   "CARRIER #01 SpareSafetyOutput(3_2)" : Bool = PLC "CARRIER #01 SpareSafetyOutput(3_2)" AT %M84.1, 1 s
   "CARRIER #01 SpareSafetyOutput(3_3)" : Bool = PLC "CARRIER #01 SpareSafetyOutput(3_3)" AT %M84.2, 1 s
   "CARRIER #01 SpareSafetyOutput(3_4)" : Bool = PLC "CARRIER #01 SpareSafetyOutput(3_4)" AT %M84.3, 1 s
   "CARRIER #01 SpareSafetyOutput(3_5)" : Bool = PLC "CARRIER #01 SpareSafetyOutput(3_5)" AT %M84.4, 1 s
   "CARRIER #01 SpareSafetyOutput(3_6)" : Bool = PLC "CARRIER #01 SpareSafetyOutput(3_6)" AT %M84.5, 1 s
   "CARRIER #01 SpareSafetyOutput(3_7)" : Bool = PLC "CARRIER #01 SpareSafetyOutput(3_7)" AT %M84.6, 1 s
   "Carrier #01_ At Command Position" : Bool = PLC DB_SDC_ERRORS_STAT.ER_AKT[49].ER_STAT[1].ERROR AT %M84.7, 1 s
   "Carrier #01_ Carrier in zone" : Int = PLC "Carrier #01_ Carrier in zone" AT %MW86, 1 s
   "Carrier #01_ Next carrier number" : Int = PLC "Carrier #01_ Next carrier number" AT %MW88, 1 s
   "Carrier 1 G120 D Status" : Bool = PLC EMS.Carrier[12].SDC_IN.DriveCommFault AT %I412.1, 1 s
   "Carrier 1 HMI Status" : Bool = PLC "Carrier 1 HMI Status" AT %I412.2, 1 s
   "Carrier 1 PnF Encoder Status" : Bool = PLC "Carrier 1 PnF Encoder Status" AT %I412.0, 1 s
   "Carrier 2  HMI Staus" : Bool = PLC "Carrier 2 HMI Status" AT %I432.2, 1 s
   "Carrier 2 G120 D Status" : Bool = PLC "Carrier 2  Drive Status" AT %I432.1, 1 s
   "Carrier 2 PnF Encoder Status" : Bool = PLC "Carrier 2 PnF Encoder Status" AT %I432.0, 1 s
   "Carrier 3  G120 D Status" : Bool = PLC "Carrier 3  Drive Status" AT %I452.1, 1 s
   "Carrier 3  PnF Encoder Status" : Bool = PLC "Carrier 3 PnF Encoder Status" AT %I452.0, 1 s
   "Carrier 3 HMI Status" : Bool = PLC "Carrier 3 HMI Status" AT %I452.2, 1 s
   "Carrier 4 G120 D Status" : Bool = PLC "Carrier 4  Drive Status" AT %I472.1, 1 s
   "Carrier 4 HMI Status" : Bool = PLC "Carrier 4 HMI Status" AT %I472.2, 1 s
   "Carrier 4 PnF Encoder Status" : Bool = PLC "Carrier 4 PnF Encoder Status" AT %I472.0, 1 s
   "Carrier_Index_HMI" : Int = PLC Carrier_Index_HMI AT %MW70, 1 s
   "Always_OFF_HMI" : Bool, internal
   "Always_ON_HMI" : Bool, internal
   "EMS_Accum_Zone_Speed" : Word = PLC EMS.AccumZnSpeed AT %DB1.DBW0, 1 s
   "PLC_IP_Address" : WString[30], internal
   "DB302_HMI_Faults_Carrier1_Faults_0" : Int = PLC DB302_HMI_Faults.Carrier1_Faults_0 AT %DB1.DBW0, 1 s
   "DB302_HMI_Faults_Carrier1_Faults_1" : Int = PLC DB302_HMI_Faults.Carrier1_Faults_1 AT %DB1.DBW0, 1 s
   "DB302_HMI_Faults_Carrier1_Faults_2" : Int = PLC DB302_HMI_Faults.Carrier1_Faults_2 AT %DB1.DBW0, 1 s
   "DB302_HMI_Faults_Carrier1_Faults_3" : Int = PLC DB302_HMI_Faults.Carrier1_Faults_3 AT %DB1.DBW0, 1 s
   "DB302_HMI_Faults_Carrier10_Faults_0" : Int = PLC DB302_HMI_Faults.Carrier10_Faults_0 AT %DB1.DBW0, 1 s
   "DB302_HMI_Faults_Carrier10_Faults_1" : Int = PLC DB302_HMI_Faults.Carrier10_Faults_1 AT %DB1.DBW0, 1 s
   "DB302_HMI_Faults_Carrier10_Faults_2" : Int = PLC DB302_HMI_Faults.Carrier10_Faults_2 AT %DB1.DBW0, 1 s
   "DB302_HMI_Faults_Carrier10_Faults_3" : Int = PLC DB302_HMI_Faults.Carrier10_Faults_3 AT %DB1.DBW0, 1 s
   "DB302_HMI_Faults_Carrier11_Faults_0" : Int = PLC DB302_HMI_Faults.Carrier11_Faults_0 AT %DB1.DBW0, 1 s
   "DB302_HMI_Faults_Carrier11_Faults_1" : Int = PLC DB302_HMI_Faults.Carrier11_Faults_1 AT %DB1.DBW0, 1 s
   "DB302_HMI_Faults_Carrier11_Faults_2" : Int = PLC DB302_HMI_Faults.Carrier11_Faults_2 AT %DB1.DBW0, 1 s
   "DB302_HMI_Faults_Carrier11_Faults_3" : Int = PLC DB302_HMI_Faults.Carrier11_Faults_3 AT %DB1.DBW0, 1 s
   "DB302_HMI_Faults_Carrier12_Faults_0" : Int = PLC DB302_HMI_Faults.Carrier12_Faults_0 AT %DB1.DBW0, 1 s
   "DB302_HMI_Faults_Carrier12_Faults_1" : Int = PLC DB302_HMI_Faults.Carrier12_Faults_1 AT %DB1.DBW0, 1 s
   "DB302_HMI_Faults_Carrier12_Faults_2" : Int = PLC DB302_HMI_Faults.Carrier12_Faults_2 AT %DB1.DBW0, 1 s
   "DB302_HMI_Faults_Carrier12_Faults_3" : Int = PLC DB302_HMI_Faults.Carrier12_Faults_3 AT %DB1.DBW0, 1 s
   "DB302_HMI_Faults_Carrier13_Faults_0" : Int = PLC DB302_HMI_Faults.Carrier13_Faults_0 AT %DB1.DBW0, 1 s
   "DB302_HMI_Faults_Carrier13_Faults_1" : Int = PLC DB302_HMI_Faults.Carrier13_Faults_1 AT %DB1.DBW0, 1 s
   "DB302_HMI_Faults_Carrier13_Faults_2" : Int = PLC DB302_HMI_Faults.Carrier13_Faults_2 AT %DB1.DBW0, 1 s
   "DB302_HMI_Faults_Carrier13_Faults_3" : Int = PLC DB302_HMI_Faults.Carrier13_Faults_3 AT %DB1.DBW0, 1 s
   "DB302_HMI_Faults_Carrier14_Faults_0" : Int = PLC DB302_HMI_Faults.Carrier14_Faults_0 AT %DB1.DBW0, 1 s
   "DB302_HMI_Faults_Carrier14_Faults_1" : Int = PLC DB302_HMI_Faults.Carrier14_Faults_1 AT %DB1.DBW0, 1 s
   "DB302_HMI_Faults_Carrier14_Faults_2" : Int = PLC DB302_HMI_Faults.Carrier14_Faults_2 AT %DB1.DBW0, 1 s
   "DB302_HMI_Faults_Carrier14_Faults_3" : Int = PLC DB302_HMI_Faults.Carrier14_Faults_3 AT %DB1.DBW0, 1 s
   "DB302_HMI_Faults_Carrier15_Faults_0" : Int = PLC DB302_HMI_Faults.Carrier15_Faults_0 AT %DB1.DBW0, 1 s
   "DB302_HMI_Faults_Carrier15_Faults_1" : Int = PLC DB302_HMI_Faults.Carrier15_Faults_1 AT %DB1.DBW0, 1 s
   "DB302_HMI_Faults_Carrier15_Faults_2" : Int = PLC DB302_HMI_Faults.Carrier15_Faults_2 AT %DB1.DBW0, 1 s
   "DB302_HMI_Faults_Carrier15_Faults_3" : Int = PLC DB302_HMI_Faults.Carrier15_Faults_3 AT %DB1.DBW0, 1 s
   "DB302_HMI_Faults_Carrier16_Faults_0" : Int = PLC DB302_HMI_Faults.Carrier16_Faults_0 AT %DB1.DBW0, 1 s
   "DB302_HMI_Faults_Carrier16_Faults_1" : Int = PLC DB302_HMI_Faults.Carrier16_Faults_1 AT %DB1.DBW0, 1 s
   "DB302_HMI_Faults_Carrier16_Faults_2" : Int = PLC DB302_HMI_Faults.Carrier16_Faults_2 AT %DB1.DBW0, 1 s
   "DB302_HMI_Faults_Carrier16_Faults_3" : Int = PLC DB302_HMI_Faults.Carrier16_Faults_3 AT %DB1.DBW0, 1 s
   "DB302_HMI_Faults_Carrier17_Faults_0" : Int = PLC DB302_HMI_Faults.Carrier17_Faults_0 AT %DB1.DBW0, 1 s
   "DB302_HMI_Faults_Carrier17_Faults_1" : Int = PLC DB302_HMI_Faults.Carrier17_Faults_1 AT %DB1.DBW0, 1 s
   "DB302_HMI_Faults_Carrier17_Faults_2" : Int = PLC DB302_HMI_Faults.Carrier17_Faults_2 AT %DB1.DBW0, 1 s
   "DB302_HMI_Faults_Carrier17_Faults_3" : Int = PLC DB302_HMI_Faults.Carrier17_Faults_3 AT %DB1.DBW0, 1 s
   "DB302_HMI_Faults_Carrier18_Faults_0" : Int = PLC DB302_HMI_Faults.Carrier18_Faults_0 AT %DB1.DBW0, 1 s
   "DB302_HMI_Faults_Carrier18_Faults_1" : Int = PLC DB302_HMI_Faults.Carrier18_Faults_1 AT %DB1.DBW0, 1 s
   "DB302_HMI_Faults_Carrier18_Faults_2" : Int = PLC DB302_HMI_Faults.Carrier18_Faults_2 AT %DB1.DBW0, 1 s
   "DB302_HMI_Faults_Carrier18_Faults_3" : Int = PLC DB302_HMI_Faults.Carrier18_Faults_3 AT %DB1.DBW0, 1 s
   "DB302_HMI_Faults_Carrier19_Faults_0" : Int = PLC DB302_HMI_Faults.Carrier19_Faults_0 AT %DB1.DBW0, 1 s
   "DB302_HMI_Faults_Carrier19_Faults_1" : Int = PLC DB302_HMI_Faults.Carrier19_Faults_1 AT %DB1.DBW0, 1 s
   "DB302_HMI_Faults_Carrier19_Faults_2" : Int = PLC DB302_HMI_Faults.Carrier19_Faults_2 AT %DB1.DBW0, 1 s
   "DB302_HMI_Faults_Carrier19_Faults_3" : Int = PLC DB302_HMI_Faults.Carrier19_Faults_3 AT %DB1.DBW0, 1 s
   "DB302_HMI_Faults_Carrier2_Faults_0" : Int = PLC DB302_HMI_Faults.Carrier2_Faults_0 AT %DB1.DBW0, 1 s
   "DB302_HMI_Faults_Carrier2_Faults_1" : Int = PLC DB302_HMI_Faults.Carrier2_Faults_1 AT %DB1.DBW0, 1 s
   "DB302_HMI_Faults_Carrier2_Faults_2" : Int = PLC DB302_HMI_Faults.Carrier2_Faults_2 AT %DB1.DBW0, 1 s
   "DB302_HMI_Faults_Carrier2_Faults_3" : Int = PLC DB302_HMI_Faults.Carrier2_Faults_3 AT %DB1.DBW0, 1 s
   "DB302_HMI_Faults_Carrier20_Faults_0" : Int = PLC DB302_HMI_Faults.Carrier20_Faults_0 AT %DB1.DBW0, 1 s
   "DB302_HMI_Faults_Carrier20_Faults_1" : Int = PLC DB302_HMI_Faults.Carrier20_Faults_1 AT %DB1.DBW0, 1 s
   "DB302_HMI_Faults_Carrier20_Faults_2" : Int = PLC DB302_HMI_Faults.Carrier20_Faults_2 AT %DB1.DBW0, 1 s
   "DB302_HMI_Faults_Carrier20_Faults_3" : Int = PLC DB302_HMI_Faults.Carrier20_Faults_3 AT %DB1.DBW0, 1 s
   "DB302_HMI_Faults_Carrier21_Faults_0" : Int = PLC DB302_HMI_Faults.Carrier21_Faults_0 AT %DB1.DBW0, 1 s
   "DB302_HMI_Faults_Carrier21_Faults_1" : Int = PLC DB302_HMI_Faults.Carrier21_Faults_1 AT %DB1.DBW0, 1 s
   "DB302_HMI_Faults_Carrier21_Faults_2" : Int = PLC DB302_HMI_Faults.Carrier21_Faults_2 AT %DB1.DBW0, 1 s
   "DB302_HMI_Faults_Carrier21_Faults_3" : Int = PLC DB302_HMI_Faults.Carrier21_Faults_3 AT %DB1.DBW0, 1 s
   "DB302_HMI_Faults_Carrier22_Faults_0" : Int = PLC DB302_HMI_Faults.Carrier22_Faults_0 AT %DB1.DBW0, 1 s
   "DB302_HMI_Faults_Carrier22_Faults_1" : Int = PLC DB302_HMI_Faults.Carrier22_Faults_1 AT %DB1.DBW0, 1 s
   "DB302_HMI_Faults_Carrier22_Faults_2" : Int = PLC DB302_HMI_Faults.Carrier22_Faults_2 AT %DB1.DBW0, 1 s
   "DB302_HMI_Faults_Carrier22_Faults_3" : Int = PLC DB302_HMI_Faults.Carrier22_Faults_3 AT %DB1.DBW0, 1 s
   "DB302_HMI_Faults_Carrier23_Faults_0" : Int = PLC DB302_HMI_Faults.Carrier23_Faults_0 AT %DB1.DBW0, 1 s
   "DB302_HMI_Faults_Carrier23_Faults_1" : Int = PLC DB302_HMI_Faults.Carrier23_Faults_1 AT %DB1.DBW0, 1 s
   "DB302_HMI_Faults_Carrier23_Faults_2" : Int = PLC DB302_HMI_Faults.Carrier23_Faults_2 AT %DB1.DBW0, 1 s
   "DB302_HMI_Faults_Carrier23_Faults_3" : Int = PLC DB302_HMI_Faults.Carrier23_Faults_3 AT %DB1.DBW0, 1 s
   "DB302_HMI_Faults_Carrier24_Faults_0" : Int = PLC DB302_HMI_Faults.Carrier24_Faults_0 AT %DB1.DBW0, 1 s
   "DB302_HMI_Faults_Carrier24_Faults_1" : Int = PLC DB302_HMI_Faults.Carrier24_Faults_1 AT %DB1.DBW0, 1 s
   "DB302_HMI_Faults_Carrier24_Faults_2" : Int = PLC DB302_HMI_Faults.Carrier24_Faults_2 AT %DB1.DBW0, 1 s
   "DB302_HMI_Faults_Carrier24_Faults_3" : Int = PLC DB302_HMI_Faults.Carrier24_Faults_3 AT %DB1.DBW0, 1 s
   "DB302_HMI_Faults_Carrier25_Faults_0" : Int = PLC DB302_HMI_Faults.Carrier25_Faults_0 AT %DB1.DBW0, 1 s
   "DB302_HMI_Faults_Carrier25_Faults_1" : Int = PLC DB302_HMI_Faults.Carrier25_Faults_1 AT %DB1.DBW0, 1 s
   "DB302_HMI_Faults_Carrier25_Faults_2" : Int = PLC DB302_HMI_Faults.Carrier25_Faults_2 AT %DB1.DBW0, 1 s
   "DB302_HMI_Faults_Carrier25_Faults_3" : Int = PLC DB302_HMI_Faults.Carrier25_Faults_3 AT %DB1.DBW0, 1 s
   "DB302_HMI_Faults_Carrier26_Faults_0" : Int = PLC DB302_HMI_Faults.Carrier26_Faults_0 AT %DB1.DBW0, 1 s
   "DB302_HMI_Faults_Carrier26_Faults_1" : Int = PLC DB302_HMI_Faults.Carrier26_Faults_1 AT %DB1.DBW0, 1 s
   "DB302_HMI_Faults_Carrier26_Faults_2" : Int = PLC DB302_HMI_Faults.Carrier26_Faults_2 AT %DB1.DBW0, 1 s
   "DB302_HMI_Faults_Carrier26_Faults_3" : Int = PLC DB302_HMI_Faults.Carrier26_Faults_3 AT %DB1.DBW0, 1 s
   "DB302_HMI_Faults_Carrier27_Faults_0" : Int = PLC DB302_HMI_Faults.Carrier27_Faults_0 AT %DB1.DBW0, 1 s
   "DB302_HMI_Faults_Carrier27_Faults_1" : Int = PLC DB302_HMI_Faults.Carrier27_Faults_1 AT %DB1.DBW0, 1 s
   "DB302_HMI_Faults_Carrier27_Faults_2" : Int = PLC DB302_HMI_Faults.Carrier27_Faults_2 AT %DB1.DBW0, 1 s
   "DB302_HMI_Faults_Carrier27_Faults_3" : Int = PLC DB302_HMI_Faults.Carrier27_Faults_3 AT %DB1.DBW0, 1 s
   "DB302_HMI_Faults_Carrier28_Faults_0" : Int = PLC DB302_HMI_Faults.Carrier28_Faults_0 AT %DB1.DBW0, 1 s
   "DB302_HMI_Faults_Carrier28_Faults_1" : Int = PLC DB302_HMI_Faults.Carrier28_Faults_1 AT %DB1.DBW0, 1 s
   "DB302_HMI_Faults_Carrier28_Faults_2" : Int = PLC DB302_HMI_Faults.Carrier28_Faults_2 AT %DB1.DBW0, 1 s
   "DB302_HMI_Faults_Carrier28_Faults_3" : Int = PLC DB302_HMI_Faults.Carrier28_Faults_3 AT %DB1.DBW0, 1 s
   "DB302_HMI_Faults_Carrier29_Faults_0" : Int = PLC DB302_HMI_Faults.Carrier29_Faults_0 AT %DB1.DBW0, 1 s
   "DB302_HMI_Faults_Carrier29_Faults_1" : Int = PLC DB302_HMI_Faults.Carrier29_Faults_1 AT %DB1.DBW0, 1 s
   "DB302_HMI_Faults_Carrier29_Faults_2" : Int = PLC DB302_HMI_Faults.Carrier29_Faults_2 AT %DB1.DBW0, 1 s
   "DB302_HMI_Faults_Carrier29_Faults_3" : Int = PLC DB302_HMI_Faults.Carrier29_Faults_3 AT %DB1.DBW0, 1 s
   "DB302_HMI_Faults_Carrier3_Faults_0" : Int = PLC DB302_HMI_Faults.Carrier3_Faults_0 AT %DB1.DBW0, 1 s
   "DB302_HMI_Faults_Carrier3_Faults_1" : Int = PLC DB302_HMI_Faults.Carrier3_Faults_1 AT %DB1.DBW0, 1 s
   "DB302_HMI_Faults_Carrier3_Faults_2" : Int = PLC DB302_HMI_Faults.Carrier3_Faults_2 AT %DB1.DBW0, 1 s
   "DB302_HMI_Faults_Carrier3_Faults_3" : Int = PLC DB302_HMI_Faults.Carrier3_Faults_3 AT %DB1.DBW0, 1 s
   "DB302_HMI_Faults_Carrier30_Faults_0" : Int = PLC DB302_HMI_Faults.Carrier30_Faults_0 AT %DB1.DBW0, 1 s
   "DB302_HMI_Faults_Carrier30_Faults_1" : Int = PLC DB302_HMI_Faults.Carrier30_Faults_1 AT %DB1.DBW0, 1 s
   "DB302_HMI_Faults_Carrier30_Faults_2" : Int = PLC DB_SDC_ERRORS_STAT.ER_AKT[16].ER_STAT[2].DRIVE_POS AT %DB1.DBW0, 1 s
   "DB302_HMI_Faults_Carrier30_Faults_3" : Int = PLC DB302_HMI_Faults.Carrier30_Faults_3 AT %DB1.DBW0, 1 s
   "DB302_HMI_Faults_Carrier31_Faults_0" : Int = PLC DB302_HMI_Faults.Carrier31_Faults_0 AT %DB1.DBW0, 1 s
   "DB302_HMI_Faults_Carrier31_Faults_1" : Int = PLC DB302_HMI_Faults.Carrier31_Faults_1 AT %DB1.DBW0, 1 s
   "DB302_HMI_Faults_Carrier31_Faults_2" : Int = PLC DB302_HMI_Faults.Carrier31_Faults_2 AT %DB1.DBW0, 1 s
   "DB302_HMI_Faults_Carrier31_Faults_3" : Int = PLC DB302_HMI_Faults.Carrier31_Faults_3 AT %DB1.DBW0, 1 s
   "DB302_HMI_Faults_Carrier32_Faults_0" : Int = PLC DB302_HMI_Faults.Carrier32_Faults_0 AT %DB1.DBW0, 1 s
   "DB302_HMI_Faults_Carrier32_Faults_1" : Int = PLC DB302_HMI_Faults.Carrier32_Faults_1 AT %DB1.DBW0, 1 s
   "DB302_HMI_Faults_Carrier32_Faults_2" : Int = PLC DB302_HMI_Faults.Carrier32_Faults_2 AT %DB1.DBW0, 1 s
   "DB302_HMI_Faults_Carrier32_Faults_3" : Int = PLC DB302_HMI_Faults.Carrier32_Faults_3 AT %DB1.DBW0, 1 s
   "DB302_HMI_Faults_Carrier33_Faults_0" : Int = PLC DB302_HMI_Faults.Carrier33_Faults_0 AT %DB1.DBW0, 1 s
   "DB302_HMI_Faults_Carrier33_Faults_1" : Int = PLC DB302_HMI_Faults.Carrier33_Faults_1 AT %DB1.DBW0, 1 s
   "DB302_HMI_Faults_Carrier33_Faults_2" : Int = PLC DB302_HMI_Faults.Carrier33_Faults_2 AT %DB1.DBW0, 1 s
   "DB302_HMI_Faults_Carrier33_Faults_3" : Int = PLC DB302_HMI_Faults.Carrier33_Faults_3 AT %DB1.DBW0, 1 s
   "DB302_HMI_Faults_Carrier34_Faults_0" : Int = PLC DB302_HMI_Faults.Carrier34_Faults_0 AT %DB1.DBW0, 1 s
   "DB302_HMI_Faults_Carrier34_Faults_1" : Int = PLC DB302_HMI_Faults.Carrier34_Faults_1 AT %DB1.DBW0, 1 s
   "DB302_HMI_Faults_Carrier34_Faults_2" : Int = PLC EMS.Carrier[23] AT %DB1.DBW0, 1 s
   "DB302_HMI_Faults_Carrier34_Faults_3" : Int = PLC DB302_HMI_Faults.Carrier34_Faults_3 AT %DB1.DBW0, 1 s
   "DB302_HMI_Faults_Carrier35_Faults_0" : Int = PLC DB302_HMI_Faults.Carrier35_Faults_0 AT %DB1.DBW0, 1 s
   "DB302_HMI_Faults_Carrier35_Faults_1" : Int = PLC DB302_HMI_Faults.Carrier35_Faults_1 AT %DB1.DBW0, 1 s
   "DB302_HMI_Faults_Carrier35_Faults_2" : Int = PLC DB302_HMI_Faults.Carrier35_Faults_2 AT %DB1.DBW0, 1 s
   "DB302_HMI_Faults_Carrier35_Faults_3" : Int = PLC DB302_HMI_Faults.Carrier35_Faults_3 AT %DB1.DBW0, 1 s
   "DB302_HMI_Faults_Carrier36_Faults_0" : Int = PLC DB302_HMI_Faults.Carrier36_Faults_0 AT %DB1.DBW0, 1 s
   "DB302_HMI_Faults_Carrier36_Faults_1" : Int = PLC DB302_HMI_Faults.Carrier36_Faults_1 AT %DB1.DBW0, 1 s
   "DB302_HMI_Faults_Carrier36_Faults_2" : Int = PLC DB302_HMI_Faults.Carrier36_Faults_2 AT %DB1.DBW0, 1 s
   "DB302_HMI_Faults_Carrier36_Faults_3" : Int = PLC DB302_HMI_Faults.Carrier36_Faults_3 AT %DB1.DBW0, 1 s
   "DB302_HMI_Faults_Carrier37_Faults_0" : Int = PLC DB302_HMI_Faults.Carrier37_Faults_0 AT %DB1.DBW0, 1 s
   "DB302_HMI_Faults_Carrier37_Faults_1" : Int = PLC DB302_HMI_Faults.Carrier37_Faults_1 AT %DB1.DBW0, 1 s
   "DB302_HMI_Faults_Carrier37_Faults_2" : Int = PLC DB302_HMI_Faults.Carrier37_Faults_2 AT %DB1.DBW0, 1 s
   "DB302_HMI_Faults_Carrier37_Faults_3" : Int = PLC DB302_HMI_Faults.Carrier37_Faults_3 AT %DB1.DBW0, 1 s
   "DB302_HMI_Faults_Carrier38_Faults_0" : Int = PLC DB302_HMI_Faults.Carrier38_Faults_0 AT %DB1.DBW0, 1 s
   "DB302_HMI_Faults_Carrier38_Faults_1" : Int = PLC DB302_HMI_Faults.Carrier38_Faults_1 AT %DB1.DBW0, 1 s
   "DB302_HMI_Faults_Carrier38_Faults_2" : Int = PLC DB302_HMI_Faults.Carrier38_Faults_2 AT %DB1.DBW0, 1 s
   "DB302_HMI_Faults_Carrier38_Faults_3" : Int = PLC DB302_HMI_Faults.Carrier38_Faults_3 AT %DB1.DBW0, 1 s
   "DB302_HMI_Faults_Carrier39_Faults_0" : Int = PLC DB302_HMI_Faults.Carrier39_Faults_0 AT %DB1.DBW0, 1 s
   "DB302_HMI_Faults_Carrier39_Faults_1" : Int = PLC DB302_HMI_Faults.Carrier39_Faults_1 AT %DB1.DBW0, 1 s
   "DB302_HMI_Faults_Carrier39_Faults_2" : Int = PLC DB302_HMI_Faults.Carrier39_Faults_2 AT %DB1.DBW0, 1 s
   "DB302_HMI_Faults_Carrier39_Faults_3" : Int = PLC DB302_HMI_Faults.Carrier39_Faults_3 AT %DB1.DBW0, 1 s
   "DB302_HMI_Faults_Carrier4_Faults_0" : Int = PLC DB302_HMI_Faults.Carrier4_Faults_0 AT %DB1.DBW0, 1 s
   "DB302_HMI_Faults_Carrier4_Faults_1" : Int = PLC DB302_HMI_Faults.Carrier4_Faults_1 AT %DB1.DBW0, 1 s
   "DB302_HMI_Faults_Carrier4_Faults_2" : Int = PLC DB302_HMI_Faults.Carrier4_Faults_2 AT %DB1.DBW0, 1 s
   "DB302_HMI_Faults_Carrier4_Faults_3" : Int = PLC DB_SDC_BARCODE_INSERTS.INSERT[10].COURSEHIGH AT %DB1.DBW0, 1 s
   "DB302_HMI_Faults_Carrier40_Faults_0" : Int = PLC DB302_HMI_Faults.Carrier40_Faults_0 AT %DB1.DBW0, 1 s
   "DB302_HMI_Faults_Carrier40_Faults_1" : Int = PLC DB302_HMI_Faults.Carrier40_Faults_1 AT %DB1.DBW0, 1 s
   "DB302_HMI_Faults_Carrier40_Faults_2" : Int = PLC DB302_HMI_Faults.Carrier40_Faults_2 AT %DB1.DBW0, 1 s
   "DB302_HMI_Faults_Carrier40_Faults_3" : Int = PLC DB302_HMI_Faults.Carrier40_Faults_3 AT %DB1.DBW0, 1 s
   "DB302_HMI_Faults_Carrier41_Faults_0" : Int = PLC DB302_HMI_Faults.Carrier41_Faults_0 AT %DB1.DBW0, 1 s
   "DB302_HMI_Faults_Carrier41_Faults_1" : Int = PLC DB302_HMI_Faults.Carrier41_Faults_1 AT %DB1.DBW0, 1 s
   "DB302_HMI_Faults_Carrier41_Faults_2" : Int = PLC DB302_HMI_Faults.Carrier41_Faults_2 AT %DB1.DBW0, 1 s
   "DB302_HMI_Faults_Carrier41_Faults_3" : Int = PLC DB302_HMI_Faults.Carrier41_Faults_3 AT %DB1.DBW0, 1 s
   "DB302_HMI_Faults_Carrier42_Faults_0" : Int = PLC DB302_HMI_Faults.Carrier42_Faults_0 AT %DB1.DBW0, 1 s
   "DB302_HMI_Faults_Carrier42_Faults_1" : Int = PLC DB302_HMI_Faults.Carrier42_Faults_1 AT %DB1.DBW0, 1 s
   "DB302_HMI_Faults_Carrier42_Faults_2" : Int = PLC DB302_HMI_Faults.Carrier42_Faults_2 AT %DB1.DBW0, 1 s
   "DB302_HMI_Faults_Carrier42_Faults_3" : Int = PLC DB302_HMI_Faults.Carrier42_Faults_3 AT %DB1.DBW0, 1 s
   "DB302_HMI_Faults_Carrier43_Faults_0" : Int = PLC DB302_HMI_Faults.Carrier43_Faults_0 AT %DB1.DBW0, 1 s
   "DB302_HMI_Faults_Carrier43_Faults_1" : Int = PLC DB302_HMI_Faults.Carrier43_Faults_1 AT %DB1.DBW0, 1 s
   "DB302_HMI_Faults_Carrier43_Faults_2" : Int = PLC DB302_HMI_Faults.Carrier43_Faults_2 AT %DB1.DBW0, 1 s
   "DB302_HMI_Faults_Carrier43_Faults_3" : Int = PLC DB302_HMI_Faults.Carrier43_Faults_3 AT %DB1.DBW0, 1 s
   "DB302_HMI_Faults_Carrier44_Faults_0" : Int = PLC DB302_HMI_Faults.Carrier44_Faults_0 AT %DB1.DBW0, 1 s
   "DB302_HMI_Faults_Carrier44_Faults_1" : Int = PLC DB302_HMI_Faults.Carrier44_Faults_1 AT %DB1.DBW0, 1 s
   "DB302_HMI_Faults_Carrier44_Faults_2" : Int = PLC DB302_HMI_Faults.Carrier44_Faults_2 AT %DB1.DBW0, 1 s
   "DB302_HMI_Faults_Carrier44_Faults_3" : Int = PLC DB302_HMI_Faults.Carrier44_Faults_3 AT %DB1.DBW0, 1 s
   "DB302_HMI_Faults_Carrier45_Faults_0" : Int = PLC DB302_HMI_Faults.Carrier45_Faults_0 AT %DB1.DBW0, 1 s
   "DB302_HMI_Faults_Carrier45_Faults_1" : Int = PLC DB302_HMI_Faults.Carrier45_Faults_1 AT %DB1.DBW0, 1 s
   "DB302_HMI_Faults_Carrier45_Faults_2" : Int = PLC DB302_HMI_Faults.Carrier45_Faults_2 AT %DB1.DBW0, 1 s
   "DB302_HMI_Faults_Carrier45_Faults_3" : Int = PLC DB302_HMI_Faults.Carrier45_Faults_3 AT %DB1.DBW0, 1 s
   "DB302_HMI_Faults_Carrier46_Faults_0" : Int = PLC DB302_HMI_Faults.Carrier46_Faults_0 AT %DB1.DBW0, 1 s
   "DB302_HMI_Faults_Carrier46_Faults_1" : Int = PLC DB302_HMI_Faults.Carrier46_Faults_1 AT %DB1.DBW0, 1 s
   "DB302_HMI_Faults_Carrier46_Faults_2" : Int = PLC DB302_HMI_Faults.Carrier46_Faults_2 AT %DB1.DBW0, 1 s
   "DB302_HMI_Faults_Carrier46_Faults_3" : Int = PLC DB302_HMI_Faults.Carrier46_Faults_3 AT %DB1.DBW0, 1 s
   "DB302_HMI_Faults_Carrier47_Faults_0" : Int = PLC DB302_HMI_Faults.Carrier47_Faults_0 AT %DB1.DBW0, 1 s
   "DB302_HMI_Faults_Carrier47_Faults_1" : Int = PLC DB302_HMI_Faults.Carrier47_Faults_1 AT %DB1.DBW0, 1 s
   "DB302_HMI_Faults_Carrier47_Faults_2" : Int = PLC DB302_HMI_Faults.Carrier47_Faults_2 AT %DB1.DBW0, 1 s
   "DB302_HMI_Faults_Carrier47_Faults_3" : Int = PLC DB302_HMI_Faults.Carrier47_Faults_3 AT %DB1.DBW0, 1 s
   "DB302_HMI_Faults_Carrier48_Faults_0" : Int = PLC DB302_HMI_Faults.Carrier48_Faults_0 AT %DB1.DBW0, 1 s
   "DB302_HMI_Faults_Carrier48_Faults_1" : Int = PLC DB302_HMI_Faults.Carrier48_Faults_1 AT %DB1.DBW0, 1 s
   "DB302_HMI_Faults_Carrier48_Faults_2" : Int = PLC DB302_HMI_Faults.Carrier48_Faults_2 AT %DB1.DBW0, 1 s
   "DB302_HMI_Faults_Carrier48_Faults_3" : Int = PLC DB302_HMI_Faults.Carrier48_Faults_3 AT %DB1.DBW0, 1 s
   "DB302_HMI_Faults_Carrier49_Faults_0" : Int = PLC DB302_HMI_Faults.Carrier49_Faults_0 AT %DB1.DBW0, 1 s
   "DB302_HMI_Faults_Carrier49_Faults_1" : Int = PLC DB302_HMI_Faults.Carrier49_Faults_1 AT %DB1.DBW0, 1 s
   "DB302_HMI_Faults_Carrier49_Faults_2" : Int = PLC DB302_HMI_Faults.Carrier49_Faults_2 AT %DB1.DBW0, 1 s
   "DB302_HMI_Faults_Carrier49_Faults_3" : Int = PLC DB302_HMI_Faults.Carrier49_Faults_3 AT %DB1.DBW0, 1 s
   "DB302_HMI_Faults_Carrier5_Faults_0" : Int = PLC DB302_HMI_Faults.Carrier5_Faults_0 AT %DB1.DBW0, 1 s
   "DB302_HMI_Faults_Carrier5_Faults_1" : Int = PLC DB302_HMI_Faults.Carrier5_Faults_1 AT %DB1.DBW0, 1 s
   "DB302_HMI_Faults_Carrier5_Faults_2" : Int = PLC DB302_HMI_Faults.Carrier5_Faults_2 AT %DB1.DBW0, 1 s
   "DB302_HMI_Faults_Carrier5_Faults_3" : Int = PLC DB302_HMI_Faults.Carrier5_Faults_3 AT %DB1.DBW0, 1 s
   "DB302_HMI_Faults_Carrier50_Faults_0" : Int = PLC DB302_HMI_Faults.Carrier50_Faults_0 AT %DB1.DBW0, 1 s
   "DB302_HMI_Faults_Carrier50_Faults_1" : Int = PLC DB302_HMI_Faults.Carrier50_Faults_1 AT %DB1.DBW0, 1 s
   "DB302_HMI_Faults_Carrier50_Faults_2" : Int = PLC DB302_HMI_Faults.Carrier50_Faults_2 AT %DB1.DBW0, 1 s
   "DB302_HMI_Faults_Carrier50_Faults_3" : Int = PLC DB302_HMI_Faults.Carrier50_Faults_3 AT %DB1.DBW0, 1 s
   "DB302_HMI_Faults_Carrier51_Faults_0" : Int = PLC DB302_HMI_Faults.Carrier51_Faults_0 AT %DB1.DBW0, 1 s
   "DB302_HMI_Faults_Carrier51_Faults_1" : Int = PLC DB302_HMI_Faults.Carrier51_Faults_1 AT %DB1.DBW0, 1 s
   "DB302_HMI_Faults_Carrier51_Faults_2" : Int = PLC DB302_HMI_Faults.Carrier51_Faults_2 AT %DB1.DBW0, 1 s
   "DB302_HMI_Faults_Carrier51_Faults_3" : Int = PLC DB302_HMI_Faults.Carrier51_Faults_3 AT %DB1.DBW0, 1 s
   "DB302_HMI_Faults_Carrier52_Faults_0" : Int = PLC DB302_HMI_Faults.Carrier52_Faults_0 AT %DB1.DBW0, 1 s
   "DB302_HMI_Faults_Carrier52_Faults_1" : Int = PLC DB302_HMI_Faults.Carrier52_Faults_1 AT %DB1.DBW0, 1 s
   "DB302_HMI_Faults_Carrier52_Faults_2" : Int = PLC DB302_HMI_Faults.Carrier52_Faults_2 AT %DB1.DBW0, 1 s
   "DB302_HMI_Faults_Carrier52_Faults_3" : Int = PLC DB_SDC_BARCODE_INSERTS.INSERT[4].INSERTLOW AT %DB1.DBW0, 1 s
   "DB302_HMI_Faults_Carrier53_Faults_0" : Int = PLC DB302_HMI_Faults.Carrier53_Faults_0 AT %DB1.DBW0, 1 s
   "DB302_HMI_Faults_Carrier53_Faults_1" : Int = PLC DB302_HMI_Faults.Carrier53_Faults_1 AT %DB1.DBW0, 1 s
   "DB302_HMI_Faults_Carrier53_Faults_2" : Int = PLC DB302_HMI_Faults.Carrier53_Faults_2 AT %DB1.DBW0, 1 s
   "DB302_HMI_Faults_Carrier53_Faults_3" : Int = PLC DB302_HMI_Faults.Carrier53_Faults_3 AT %DB1.DBW0, 1 s
   "DB302_HMI_Faults_Carrier54_Faults_0" : Int = PLC DB302_HMI_Faults.Carrier54_Faults_0 AT %DB1.DBW0, 1 s
   "DB302_HMI_Faults_Carrier54_Faults_1" : Int = PLC DB302_HMI_Faults.Carrier54_Faults_1 AT %DB1.DBW0, 1 s
   "DB302_HMI_Faults_Carrier54_Faults_2" : Int = PLC DB302_HMI_Faults.Carrier54_Faults_2 AT %DB1.DBW0, 1 s
   "DB302_HMI_Faults_Carrier54_Faults_3" : Int = PLC DB302_HMI_Faults.Carrier54_Faults_3 AT %DB1.DBW0, 1 s
   "DB302_HMI_Faults_Carrier55_Faults_0" : Int = PLC DB302_HMI_Faults.Carrier55_Faults_0 AT %DB1.DBW0, 1 s
   "DB302_HMI_Faults_Carrier55_Faults_1" : Int = PLC DB302_HMI_Faults.Carrier55_Faults_1 AT %DB1.DBW0, 1 s
   "DB302_HMI_Faults_Carrier55_Faults_2" : Int = PLC DB302_HMI_Faults.Carrier55_Faults_2 AT %DB1.DBW0, 1 s
   "DB302_HMI_Faults_Carrier55_Faults_3" : Int = PLC DB302_HMI_Faults.Carrier55_Faults_3 AT %DB1.DBW0, 1 s
   "DB302_HMI_Faults_Carrier56_Faults_0" : Int = PLC DB302_HMI_Faults.Carrier56_Faults_0 AT %DB1.DBW0, 1 s
   "DB302_HMI_Faults_Carrier56_Faults_1" : Int = PLC DB302_HMI_Faults.Carrier56_Faults_1 AT %DB1.DBW0, 1 s
   "DB302_HMI_Faults_Carrier56_Faults_2" : Int = PLC DB302_HMI_Faults.Carrier56_Faults_2 AT %DB1.DBW0, 1 s
   "DB302_HMI_Faults_Carrier56_Faults_3" : Int = PLC DB302_HMI_Faults.Carrier56_Faults_3 AT %DB1.DBW0, 1 s
   "DB302_HMI_Faults_Carrier57_Faults_0" : Int = PLC DB302_HMI_Faults.Carrier57_Faults_0 AT %DB1.DBW0, 1 s
   "DB302_HMI_Faults_Carrier57_Faults_1" : Int = PLC DB302_HMI_Faults.Carrier57_Faults_1 AT %DB1.DBW0, 1 s
   "DB302_HMI_Faults_Carrier57_Faults_2" : Int = PLC DB302_HMI_Faults.Carrier57_Faults_2 AT %DB1.DBW0, 1 s
   "DB302_HMI_Faults_Carrier57_Faults_3" : Int = PLC DB302_HMI_Faults.Carrier57_Faults_3 AT %DB1.DBW0, 1 s
   "DB302_HMI_Faults_Carrier58_Faults_0" : Int = PLC DB302_HMI_Faults.Carrier58_Faults_0 AT %DB1.DBW0, 1 s
   "DB302_HMI_Faults_Carrier58_Faults_1" : Int = PLC DB302_HMI_Faults.Carrier58_Faults_1 AT %DB1.DBW0, 1 s
   "DB302_HMI_Faults_Carrier58_Faults_2" : Int = PLC DB302_HMI_Faults.Carrier58_Faults_2 AT %DB1.DBW0, 1 s
   "DB302_HMI_Faults_Carrier58_Faults_3" : Int = PLC DB302_HMI_Faults.Carrier58_Faults_3 AT %DB1.DBW0, 1 s
   "DB302_HMI_Faults_Carrier59_Faults_0" : Int = PLC DB302_HMI_Faults.Carrier59_Faults_0 AT %DB1.DBW0, 1 s
   "DB302_HMI_Faults_Carrier59_Faults_1" : Int = PLC DB302_HMI_Faults.Carrier59_Faults_1 AT %DB1.DBW0, 1 s
   "DB302_HMI_Faults_Carrier59_Faults_2" : Int = PLC DB302_HMI_Faults.Carrier59_Faults_2 AT %DB1.DBW0, 1 s
   "DB302_HMI_Faults_Carrier59_Faults_3" : Int = PLC DB302_HMI_Faults.Carrier59_Faults_3 AT %DB1.DBW0, 1 s
   "DB302_HMI_Faults_Carrier6_Faults_0" : Int = PLC DB302_HMI_Faults.Carrier6_Faults_0 AT %DB1.DBW0, 1 s
   "DB302_HMI_Faults_Carrier6_Faults_1" : Int = PLC DB302_HMI_Faults.Carrier6_Faults_1 AT %DB1.DBW0, 1 s
   "DB302_HMI_Faults_Carrier6_Faults_2" : Int = PLC DB302_HMI_Faults.Carrier6_Faults_2 AT %DB1.DBW0, 1 s
   "DB302_HMI_Faults_Carrier6_Faults_3" : Int = PLC DB302_HMI_Faults.Carrier6_Faults_3 AT %DB1.DBW0, 1 s
   "DB302_HMI_Faults_Carrier60_Faults_0" : Int = PLC DB302_HMI_Faults.Carrier60_Faults_0 AT %DB1.DBW0, 1 s
   "DB302_HMI_Faults_Carrier60_Faults_1" : Int = PLC DB302_HMI_Faults.Carrier60_Faults_1 AT %DB1.DBW0, 1 s
   "DB302_HMI_Faults_Carrier60_Faults_2" : Int = PLC DB302_HMI_Faults.Carrier60_Faults_2 AT %DB1.DBW0, 1 s
   "DB302_HMI_Faults_Carrier60_Faults_3" : Int = PLC DB302_HMI_Faults.Carrier60_Faults_3 AT %DB1.DBW0, 1 s
   "DB302_HMI_Faults_Carrier61_Faults_0" : Int = PLC DB302_HMI_Faults.Carrier61_Faults_0 AT %DB1.DBW0, 1 s
   "DB302_HMI_Faults_Carrier61_Faults_1" : Int = PLC DB302_HMI_Faults.Carrier61_Faults_1 AT %DB1.DBW0, 1 s
   "DB302_HMI_Faults_Carrier61_Faults_2" : Int = PLC DB302_HMI_Faults.Carrier61_Faults_2 AT %DB1.DBW0, 1 s
   "DB302_HMI_Faults_Carrier61_Faults_3" : Int = PLC DB302_HMI_Faults.Carrier61_Faults_3 AT %DB1.DBW0, 1 s
   "DB302_HMI_Faults_Carrier62_Faults_0" : Int = PLC DB302_HMI_Faults.Carrier62_Faults_0 AT %DB1.DBW0, 1 s
   "DB302_HMI_Faults_Carrier62_Faults_1" : Int = PLC DB302_HMI_Faults.Carrier62_Faults_1 AT %DB1.DBW0, 1 s
   "DB302_HMI_Faults_Carrier62_Faults_2" : Int = PLC DB302_HMI_Faults.Carrier62_Faults_2 AT %DB1.DBW0, 1 s
   "DB302_HMI_Faults_Carrier62_Faults_3" : Int = PLC DB302_HMI_Faults.Carrier62_Faults_3 AT %DB1.DBW0, 1 s
   "DB302_HMI_Faults_Carrier63_Faults_0" : Int = PLC DB302_HMI_Faults.Carrier63_Faults_0 AT %DB1.DBW0, 1 s
   "DB302_HMI_Faults_Carrier63_Faults_1" : Int = PLC DB302_HMI_Faults.Carrier63_Faults_1 AT %DB1.DBW0, 1 s
   "DB302_HMI_Faults_Carrier63_Faults_2" : Int = PLC DB302_HMI_Faults.Carrier63_Faults_2 AT %DB1.DBW0, 1 s
   "DB302_HMI_Faults_Carrier63_Faults_3" : Int = PLC DB302_HMI_Faults.Carrier63_Faults_3 AT %DB1.DBW0, 1 s
   "DB302_HMI_Faults_Carrier64_Faults_0" : Int = PLC DB302_HMI_Faults.Carrier64_Faults_0 AT %DB1.DBW0, 1 s
   "DB302_HMI_Faults_Carrier64_Faults_1" : Int = PLC DB302_HMI_Faults.Carrier64_Faults_1 AT %DB1.DBW0, 1 s
   "DB302_HMI_Faults_Carrier64_Faults_2" : Int = PLC DB302_HMI_Faults.Carrier64_Faults_2 AT %DB1.DBW0, 1 s
   "DB302_HMI_Faults_Carrier64_Faults_3" : Int = PLC DB302_HMI_Faults.Carrier64_Faults_3 AT %DB1.DBW0, 1 s
   "DB302_HMI_Faults_Carrier65_Faults_0" : Int = PLC DB302_HMI_Faults.Carrier65_Faults_0 AT %DB1.DBW0, 1 s
   "DB302_HMI_Faults_Carrier65_Faults_1" : Int = PLC DB302_HMI_Faults.Carrier65_Faults_1 AT %DB1.DBW0, 1 s
   "DB302_HMI_Faults_Carrier65_Faults_2" : Int = PLC DB302_HMI_Faults.Carrier65_Faults_2 AT %DB1.DBW0, 1 s
   "DB302_HMI_Faults_Carrier65_Faults_3" : Int = PLC DB302_HMI_Faults.Carrier65_Faults_3 AT %DB1.DBW0, 1 s
   "DB302_HMI_Faults_Carrier66_Faults_0" : Int = PLC DB302_HMI_Faults.Carrier66_Faults_0 AT %DB1.DBW0, 1 s
   "DB302_HMI_Faults_Carrier66_Faults_1" : Int = PLC DB302_HMI_Faults.Carrier66_Faults_1 AT %DB1.DBW0, 1 s
   "DB302_HMI_Faults_Carrier66_Faults_2" : Int = PLC DB302_HMI_Faults.Carrier66_Faults_2 AT %DB1.DBW0, 1 s
   "DB302_HMI_Faults_Carrier66_Faults_3" : Int = PLC DB302_HMI_Faults.Carrier66_Faults_3 AT %DB1.DBW0, 1 s
   "DB302_HMI_Faults_Carrier67_Faults_0" : Int = PLC DB302_HMI_Faults.Carrier67_Faults_0 AT %DB1.DBW0, 1 s
   "DB302_HMI_Faults_Carrier67_Faults_1" : Int = PLC DB302_HMI_Faults.Carrier67_Faults_1 AT %DB1.DBW0, 1 s
   "DB302_HMI_Faults_Carrier67_Faults_2" : Int = PLC DB302_HMI_Faults.Carrier67_Faults_2 AT %DB1.DBW0, 1 s
   "DB302_HMI_Faults_Carrier67_Faults_3" : Int = PLC DB302_HMI_Faults.Carrier67_Faults_3 AT %DB1.DBW0, 1 s
   "DB302_HMI_Faults_Carrier68_Faults_0" : Int = PLC DB302_HMI_Faults.Carrier68_Faults_0 AT %DB1.DBW0, 1 s
   "DB302_HMI_Faults_Carrier68_Faults_1" : Int = PLC DB302_HMI_Faults.Carrier68_Faults_1 AT %DB1.DBW0, 1 s
   "DB302_HMI_Faults_Carrier68_Faults_2" : Int = PLC DB302_HMI_Faults.Carrier68_Faults_2 AT %DB1.DBW0, 1 s
   "DB302_HMI_Faults_Carrier68_Faults_3" : Int = PLC DB302_HMI_Faults.Carrier68_Faults_3 AT %DB1.DBW0, 1 s
   "DB302_HMI_Faults_Carrier69_Faults_0" : Int = PLC DB302_HMI_Faults.Carrier69_Faults_0 AT %DB1.DBW0, 1 s
   "DB302_HMI_Faults_Carrier69_Faults_1" : Int = PLC DB302_HMI_Faults.Carrier69_Faults_1 AT %DB1.DBW0, 1 s
   "DB302_HMI_Faults_Carrier69_Faults_2" : Int = PLC DB302_HMI_Faults.Carrier69_Faults_2 AT %DB1.DBW0, 1 s
   "DB302_HMI_Faults_Carrier69_Faults_3" : Int = PLC DB302_HMI_Faults.Carrier69_Faults_3 AT %DB1.DBW0, 1 s
   "DB302_HMI_Faults_Carrier7_Faults_0" : Int = PLC DB302_HMI_Faults.Carrier7_Faults_0 AT %DB1.DBW0, 1 s
   "DB302_HMI_Faults_Carrier7_Faults_1" : Int = PLC DB302_HMI_Faults.Carrier7_Faults_1 AT %DB1.DBW0, 1 s
   "DB302_HMI_Faults_Carrier7_Faults_2" : Int = PLC DB302_HMI_Faults.Carrier7_Faults_2 AT %DB1.DBW0, 1 s
   "DB302_HMI_Faults_Carrier7_Faults_3" : Int = PLC DB302_HMI_Faults.Carrier7_Faults_3 AT %DB1.DBW0, 1 s
   "DB302_HMI_Faults_Carrier70_Faults_0" : Int = PLC DB302_HMI_Faults.Carrier70_Faults_0 AT %DB1.DBW0, 1 s
   "DB302_HMI_Faults_Carrier70_Faults_1" : Int = PLC DB302_HMI_Faults.Carrier70_Faults_1 AT %DB1.DBW0, 1 s
   "DB302_HMI_Faults_Carrier70_Faults_2" : Int = PLC DB302_HMI_Faults.Carrier70_Faults_2 AT %DB1.DBW0, 1 s
   "DB302_HMI_Faults_Carrier70_Faults_3" : Int = PLC DB302_HMI_Faults.Carrier70_Faults_3 AT %DB1.DBW0, 1 s
   "DB302_HMI_Faults_Carrier71_Faults_0" : Int = PLC DB302_HMI_Faults.Carrier71_Faults_0 AT %DB1.DBW0, 1 s